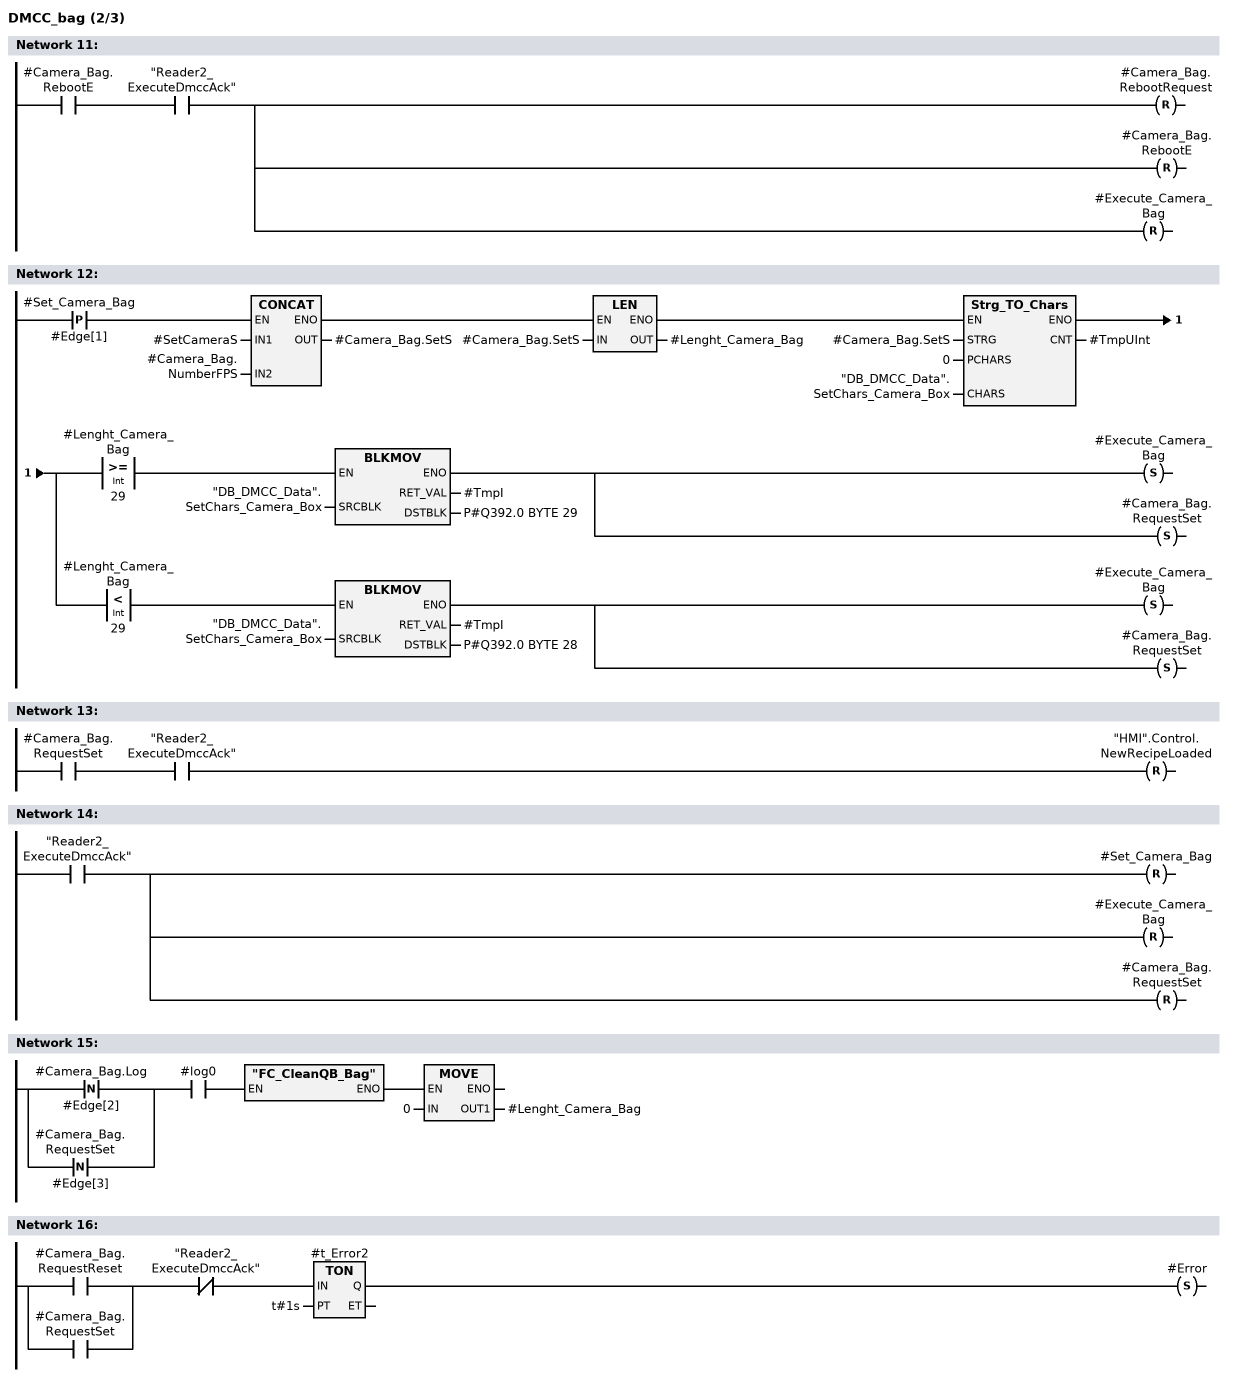
   RUNG wire#powerrail
      Contact( #Camera_Bag.RebootE )
      Contact( "Reader2_ExecuteDmccAck" )
      wire#w1
      R_Coil( #Camera_Bag.RebootRequest )
   END_RUNG
   RUNG wire#w1
      R_Coil( #Camera_Bag.RebootE )
   END_RUNG
   RUNG wire#w1
      R_Coil( #Execute_Camera_Bag )
   END_RUNG
   // the same network as SCL:
   IF #Camera_Bag.RebootE AND "Reader2_ExecuteDmccAck" THEN #Camera_Bag.RebootRequest := FALSE; END_IF;
   #_w1 := #Camera_Bag.RebootE AND "Reader2_ExecuteDmccAck";
   IF #_w1 THEN
       #Camera_Bag.RebootE := FALSE;
       #Execute_Camera_Bag := FALSE;
   END_IF;
END_REGION

REGION Network 12
   // no SCL statement known for Strg_TO_Chars: written as a call
   // ENO of a box is taken as its EN; it also drops when the box reports an error
   #_w1 := #Set_Camera_Bag AND NOT #Edge[1];   // rising edge of #Set_Camera_Bag
   #Edge[1] := #Set_Camera_Bag;
   IF #_w1 THEN
       #Camera_Bag.SetS := CONCAT(IN1 := #SetCameraS, IN2 := #Camera_Bag.NumberFPS);
       #Lenght_Camera_Bag := LEN(IN := #Camera_Bag.SetS);
       Strg_TO_Chars(Strg := #Camera_Bag.SetS,
                     pChars := 0,
                     Chars := "DB_DMCC_Data".SetChars_Camera_Box,
                     Cnt => #TmpUInt);
   END_IF;
   IF #_w1 AND (#Lenght_Camera_Bag >= 29) THEN
       #TmpI := BLKMOV(SRCBLK := "DB_DMCC_Data".SetChars_Camera_Box, DSTBLK => P#Q392.0 BYTE 29);
       #Execute_Camera_Bag := TRUE;
       #Camera_Bag.RequestSet := TRUE;
   END_IF;
   IF #_w1 AND (#Lenght_Camera_Bag < 29) THEN
       #TmpI := BLKMOV(SRCBLK := "DB_DMCC_Data".SetChars_Camera_Box, DSTBLK => P#Q392.0 BYTE 28);
       #Execute_Camera_Bag := TRUE;
       #Camera_Bag.RequestSet := TRUE;
   END_IF;
END_REGION

REGION Network 13
   RUNG wire#powerrail
      Contact( #Camera_Bag.RequestSet )
      Contact( "Reader2_ExecuteDmccAck" )
      R_Coil( "HMI".Control.NewRecipeLoaded )
   END_RUNG
   // the same network as SCL:
   IF #Camera_Bag.RequestSet AND "Reader2_ExecuteDmccAck" THEN
       "HMI".Control.NewRecipeLoaded := FALSE;
   END_IF;
END_REGION

REGION Network 14
   RUNG wire#powerrail
      Contact( "Reader2_ExecuteDmccAck" )
      wire#w1
      R_Coil( #Set_Camera_Bag )
   END_RUNG
   RUNG wire#w1
      R_Coil( #Execute_Camera_Bag )
   END_RUNG
   RUNG wire#w1
      R_Coil( #Camera_Bag.RequestSet )
   END_RUNG
   // the same network as SCL:
   IF "Reader2_ExecuteDmccAck" THEN
       #Set_Camera_Bag := FALSE;
       #Execute_Camera_Bag := FALSE;
       #Camera_Bag.RequestSet := FALSE;
   END_IF;
END_REGION

REGION Network 15
   RUNG wire#powerrail
      N_Contact(operand := #Camera_Bag.Log, bit := #Edge[2])
      wire#w1
      Contact( #log0 )
      "FC_CleanQB_Bag"()
      Move(in := 0, out1 => #Lenght_Camera_Bag)
   END_RUNG
   RUNG wire#powerrail
      N_Contact(operand := #Camera_Bag.RequestSet, bit := #Edge[3])
   END_RUNG wire#w1
   // the same network as SCL:
   #_w1 := NOT #Camera_Bag.Log AND #Edge[2];   // falling edge of #Camera_Bag.Log
   #Edge[2] := #Camera_Bag.Log;
   #_w2 := NOT #Camera_Bag.RequestSet AND #Edge[3];   // falling edge of #Camera_Bag.RequestSet
   #Edge[3] := #Camera_Bag.RequestSet;
   "FC_CleanQB_Bag"(EN := (#_w1 OR #_w2) AND #log0, ENO => #_w3);
   IF #_w3 THEN #Lenght_Camera_Bag := 0; END_IF;
END_REGION

REGION Network 16
   #t_Error2(IN := (#Camera_Bag.RequestReset OR #Camera_Bag.RequestSet) AND NOT "Reader2_ExecuteDmccAck",   // TON
             PT := t#1s);
   IF #t_Error2.Q THEN #Error := TRUE; END_IF;
END_REGION

REGION Network 17
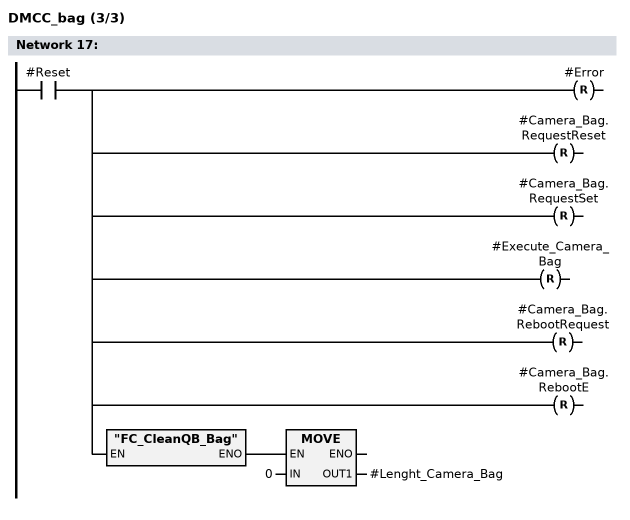
   RUNG wire#powerrail
      Contact( #Reset )
      wire#w1
      R_Coil( #Error )
   END_RUNG
   RUNG wire#w1
      R_Coil( #Camera_Bag.RequestReset )
   END_RUNG
   RUNG wire#w1
      R_Coil( #Camera_Bag.RequestSet )
   END_RUNG
   RUNG wire#w1
      R_Coil( #Execute_Camera_Bag )
   END_RUNG
   RUNG wire#w1
      R_Coil( #Camera_Bag.RebootRequest )
   END_RUNG
   RUNG wire#w1
      R_Coil( #Camera_Bag.RebootE )
   END_RUNG
   RUNG wire#w1
      "FC_CleanQB_Bag"()
      Move(in := 0, out1 => #Lenght_Camera_Bag)
   END_RUNG
   // the same network as SCL:
   IF #Reset THEN
       #Error := FALSE;
       #Camera_Bag.RequestReset := FALSE;
       #Camera_Bag.RequestSet := FALSE;
       #Execute_Camera_Bag := FALSE;
       #Camera_Bag.RebootRequest := FALSE;
       #Camera_Bag.RebootE := FALSE;
   END_IF;
   "FC_CleanQB_Bag"(EN := #Reset, ENO => #_w1);
   IF #_w1 THEN #Lenght_Camera_Bag := 0; END_IF;
END_REGION
END_FUNCTION_BLOCK

FUNCTION_BLOCK "CodeHandle"   // FB105, LAD
{ S7_Optimized_Access := 'TRUE' }
VERSION : 0.1
   VAR_INPUT
      RawCode : Array[0..86] of Char;
      Charakter : String;
      ResultLength : Int;
      Reset_faults : Bool;
      Cam_Box_Read : Bool;
   END_VAR
   VAR_OUTPUT
      LongCode_Out : String[80];
      ShortCode_Out : String[9];
      Read_BOX_EM : Bool;
      Only_ENIGMA : Bool;
      Only_MIRAI : Bool;
   END_VAR
   VAR
      Edge : Array[0..15] of Bool;
      Log1 : Bool;
      Log0 : Bool;
      CharakterPosition : Int;
      RawS : String;
      LongCode : Struct
         Long : String[80];
         Long_Part1 : String[16];
         Long_Part2 : String[12];
         Long_Part3 : String[12];
         Long_Part4 : String[16];
         Long_Part5 : String[8];
         Long_Part6 : String[8];
      END_STRUCT;
      ShortCode : Struct
         ShortCode : String[9];
      END_STRUCT;
      Enigma : TON_TIME;
   END_VAR
   VAR_TEMP
      tmp_w : Word;
      tmp_s : String;
      tmp_small : Bool;
      tmp_big : Bool;
      tmp_read : Bool;
      tmp_read_all : Bool;
   END_VAR
   VAR CONSTANT
      NoCode_ENIGMA : String := 'XXXXXXXXXXXXX';
      NoCode_MIRAI : String := 'XXXXXXXXXXXXXXXXXXXXXXXXXXXXXXXXXXXXXXXXXXXXXXXXXXXXXXXXXXXXXXXXXXXXXX';
   END_VAR
   VAR_TEMP   // added for the SCL form of the ladder/FBD networks
      _w1 : Bool;
      _w2 : Bool;
      _w3 : Bool;
      _w4 : Bool;
      _w5 : Bool;
   END_VAR
BEGIN

REGION Network 1
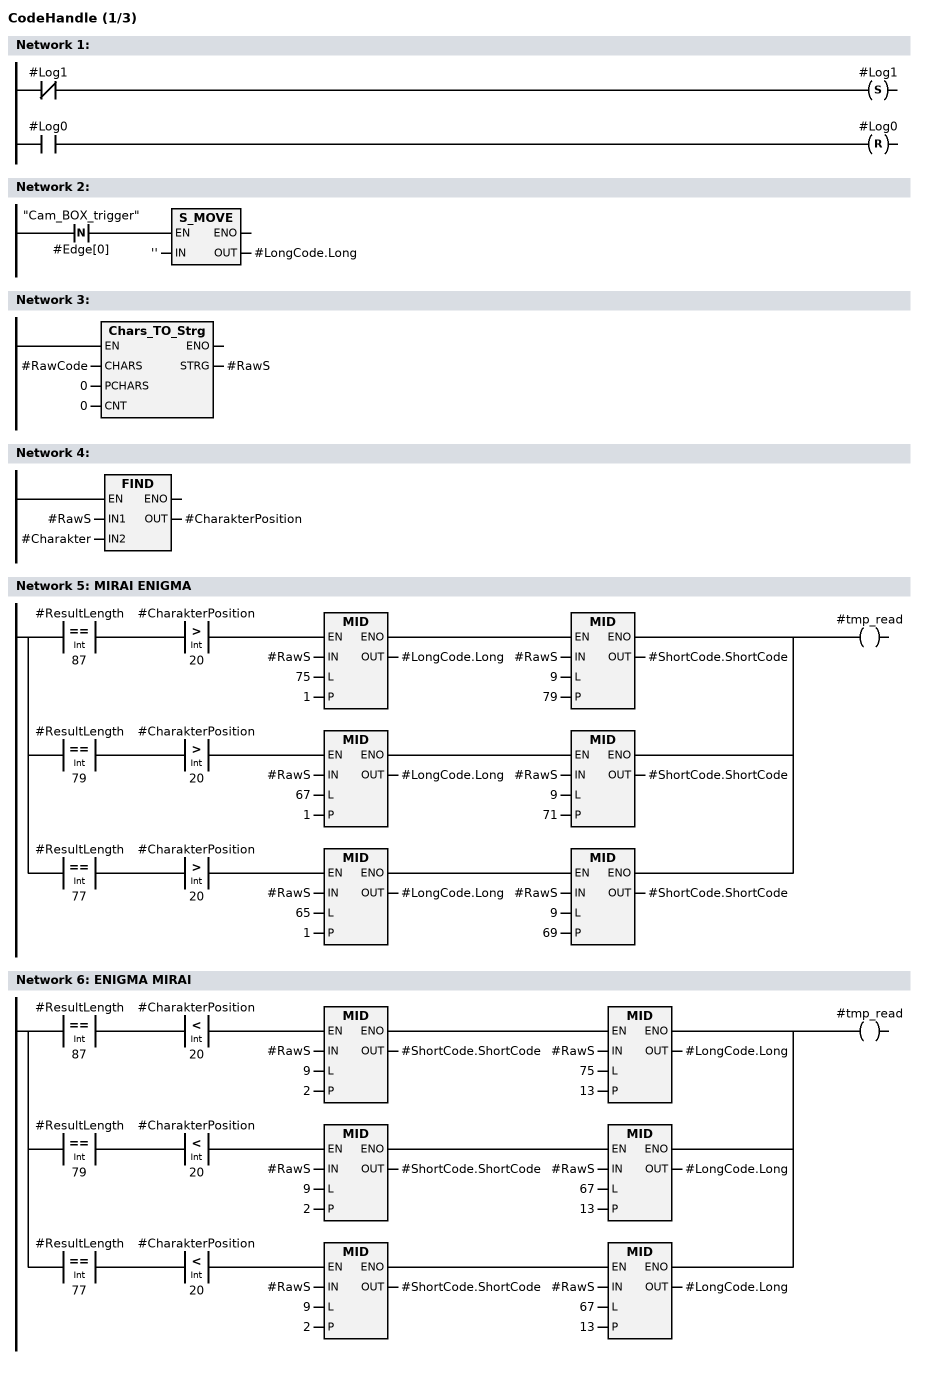
   RUNG wire#powerrail
      I_Contact( #Log1 )
      S_Coil( #Log1 )
   END_RUNG
   RUNG wire#powerrail
      Contact( #Log0 )
      R_Coil( #Log0 )
   END_RUNG
   // the same network as SCL:
   IF NOT #Log1 THEN #Log1 := TRUE; END_IF;
   IF #Log0 THEN #Log0 := FALSE; END_IF;
END_REGION

REGION Network 2
   RUNG wire#powerrail
      N_Contact(operand := "Cam_BOX_trigger", bit := #Edge[0])
      S_Move(in := '', out => #LongCode.Long)
   END_RUNG
   // the same network as SCL:
   #_w1 := NOT "Cam_BOX_trigger" AND #Edge[0];   // falling edge of "Cam_BOX_trigger"
   #Edge[0] := "Cam_BOX_trigger";
   IF #_w1 THEN #LongCode.Long := ''; END_IF;
END_REGION

REGION Network 3
   // no SCL statement known for Chars_TO_Strg: written as a call
   Chars_TO_Strg(Chars := #RawCode, pChars := 0, Cnt := 0, Strg => #RawS);
END_REGION

REGION Network 4
   #CharakterPosition := FIND(IN1 := #RawS, IN2 := #Charakter);
END_REGION

REGION Network 5: MIRAI ENIGMA
   #_w1 := (#ResultLength = 87) AND (#CharakterPosition > 20);
   IF #_w1 THEN
       #LongCode.Long := MID(IN := #RawS, L := 75, P := 1);
       #ShortCode.ShortCode := MID(IN := #RawS, L := 9, P := 79);
   END_IF;
   #_w2 := (#ResultLength = 79) AND (#CharakterPosition > 20);
   IF #_w2 THEN
       #LongCode.Long := MID(IN := #RawS, L := 67, P := 1);
       #ShortCode.ShortCode := MID(IN := #RawS, L := 9, P := 71);
   END_IF;
   #_w3 := (#ResultLength = 77) AND (#CharakterPosition > 20);
   IF #_w3 THEN
       #LongCode.Long := MID(IN := #RawS, L := 65, P := 1);
       #ShortCode.ShortCode := MID(IN := #RawS, L := 9, P := 69);
   END_IF;
   #tmp_read := #_w1 OR #_w2 OR #_w3;
END_REGION

REGION Network 6: ENIGMA MIRAI
   #_w1 := (#ResultLength = 87) AND (#CharakterPosition < 20);
   IF #_w1 THEN
       #ShortCode.ShortCode := MID(IN := #RawS, L := 9, P := 2);
       #LongCode.Long := MID(IN := #RawS, L := 75, P := 13);
   END_IF;
   #_w2 := (#ResultLength = 79) AND (#CharakterPosition < 20);
   IF #_w2 THEN
       #ShortCode.ShortCode := MID(IN := #RawS, L := 9, P := 2);
       #LongCode.Long := MID(IN := #RawS, L := 67, P := 13);
   END_IF;
   #_w3 := (#ResultLength = 77) AND (#CharakterPosition < 20);
   IF #_w3 THEN
       #ShortCode.ShortCode := MID(IN := #RawS, L := 9, P := 2);
       #LongCode.Long := MID(IN := #RawS, L := 67, P := 13);
   END_IF;
   #tmp_read := #_w1 OR #_w2 OR #_w3;
END_REGION

REGION Network 7
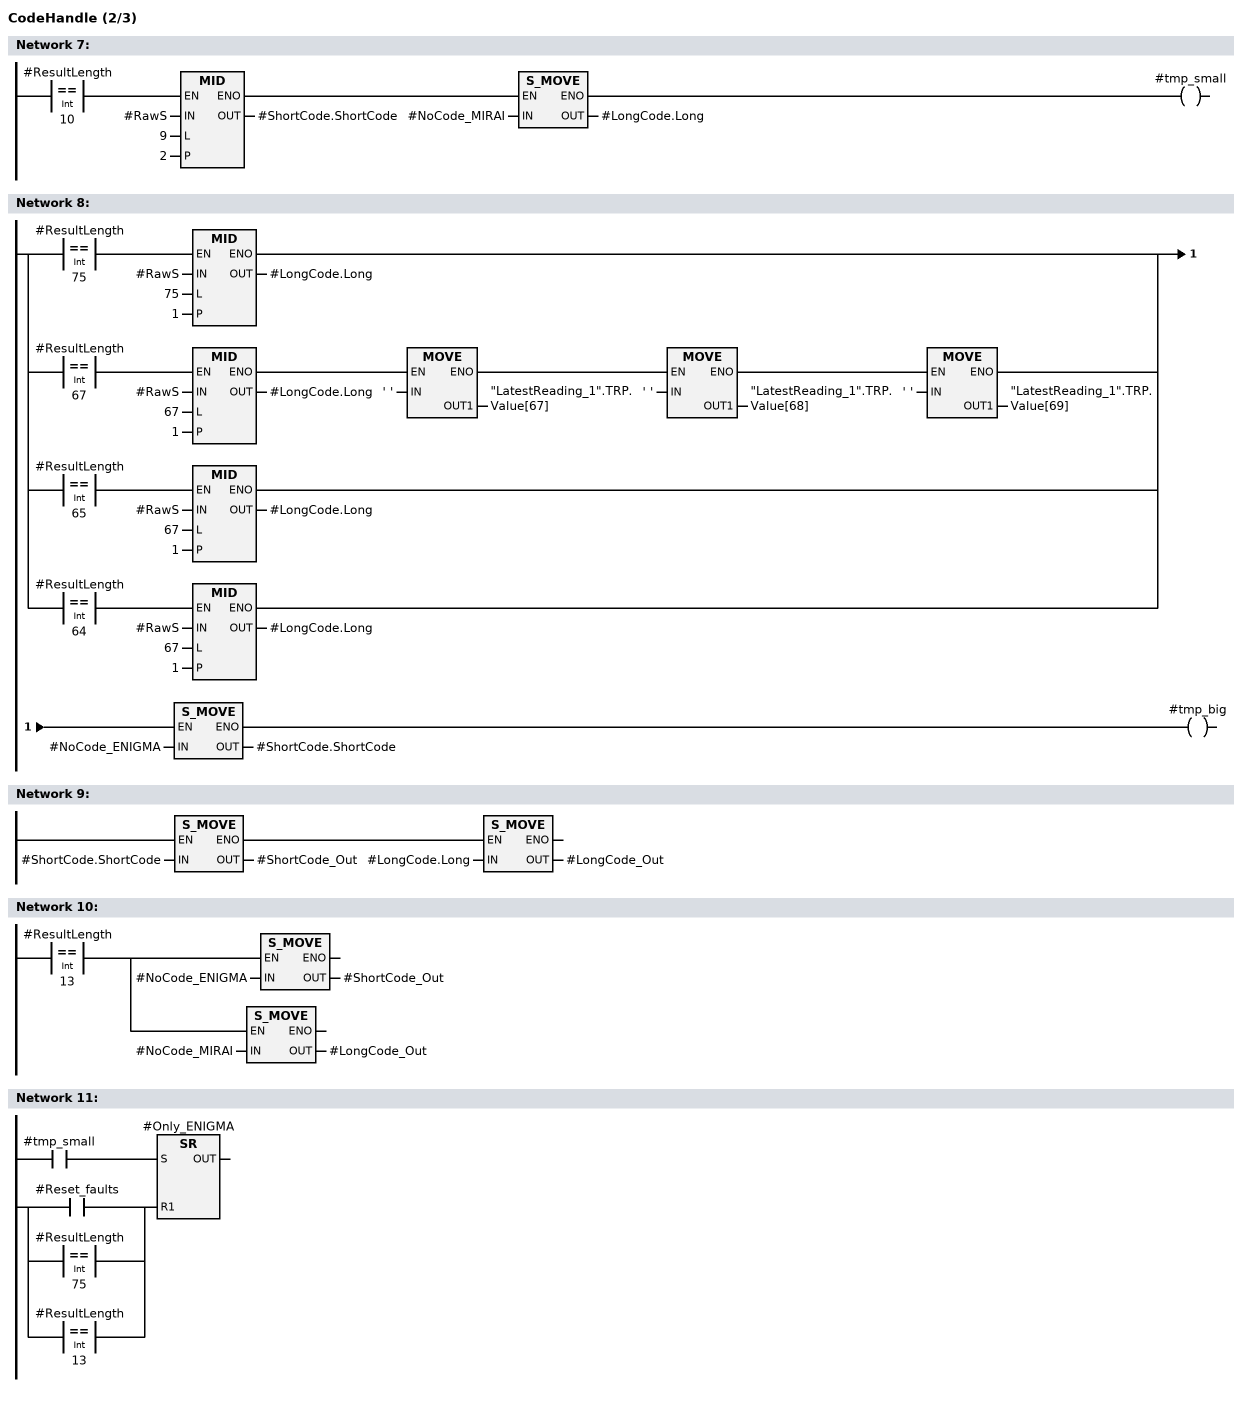
   #_w1 := #ResultLength = 10;
   IF #_w1 THEN
       #ShortCode.ShortCode := MID(IN := #RawS, L := 9, P := 2);
       #LongCode.Long := #NoCode_MIRAI;
   END_IF;
   #tmp_small := #_w1;
END_REGION

REGION Network 8
   #_w1 := #ResultLength = 75;
   IF #_w1 THEN #LongCode.Long := MID(IN := #RawS, L := 75, P := 1); END_IF;
   #_w2 := #ResultLength = 67;
   IF #_w2 THEN
       #LongCode.Long := MID(IN := #RawS, L := 67, P := 1);
       "LatestReading_1".TRP.Value[67] := ' ';
       "LatestReading_1".TRP.Value[68] := ' ';
       "LatestReading_1".TRP.Value[69] := ' ';
   END_IF;
   #_w3 := #ResultLength = 65;
   IF #_w3 THEN #LongCode.Long := MID(IN := #RawS, L := 67, P := 1); END_IF;
   #_w4 := #ResultLength = 64;
   IF #_w4 THEN #LongCode.Long := MID(IN := #RawS, L := 67, P := 1); END_IF;
   #_w5 := #_w1 OR #_w2 OR #_w3 OR #_w4;
   IF #_w5 THEN #ShortCode.ShortCode := #NoCode_ENIGMA; END_IF;
   #tmp_big := #_w5;
END_REGION

REGION Network 9
   RUNG wire#powerrail
      S_Move(in := #ShortCode.ShortCode, out => #ShortCode_Out)
      S_Move(in := #LongCode.Long, out => #LongCode_Out)
   END_RUNG
   // the same network as SCL:
   #ShortCode_Out := #ShortCode.ShortCode;
   #LongCode_Out := #LongCode.Long;
END_REGION

REGION Network 10
   RUNG wire#powerrail
      { S7_Templates := "SrcType := Int" } EQ_Contact(in1 := #ResultLength, in2 := 13)
      wire#w1
      S_Move(in := #NoCode_ENIGMA, out => #ShortCode_Out)
   END_RUNG
   RUNG wire#w1
      S_Move(in := #NoCode_MIRAI, out => #LongCode_Out)
   END_RUNG
   // the same network as SCL:
   IF #ResultLength = 13 THEN
       #ShortCode_Out := #NoCode_ENIGMA;
       #LongCode_Out := #NoCode_MIRAI;
   END_IF;
END_REGION

REGION Network 11
   RUNG wire#powerrail
      Contact( #tmp_small )
      S_SR(operand := #Only_ENIGMA, r1 := wire#w1)
   END_RUNG
   RUNG wire#powerrail
      Contact( #Reset_faults )
   END_RUNG wire#w1
   RUNG wire#powerrail
      { S7_Templates := "SrcType := Int" } EQ_Contact(in1 := #ResultLength, in2 := 75)
   END_RUNG wire#w1
   RUNG wire#powerrail
      { S7_Templates := "SrcType := Int" } EQ_Contact(in1 := #ResultLength, in2 := 13)
   END_RUNG wire#w1
   // the same network as SCL:
   IF #tmp_small THEN
       #Only_ENIGMA := TRUE;   // SR flip-flop
   END_IF;
   IF #Reset_faults OR (#ResultLength = 75) OR (#ResultLength = 13) THEN #Only_ENIGMA := FALSE; END_IF;
END_REGION

REGION Network 12
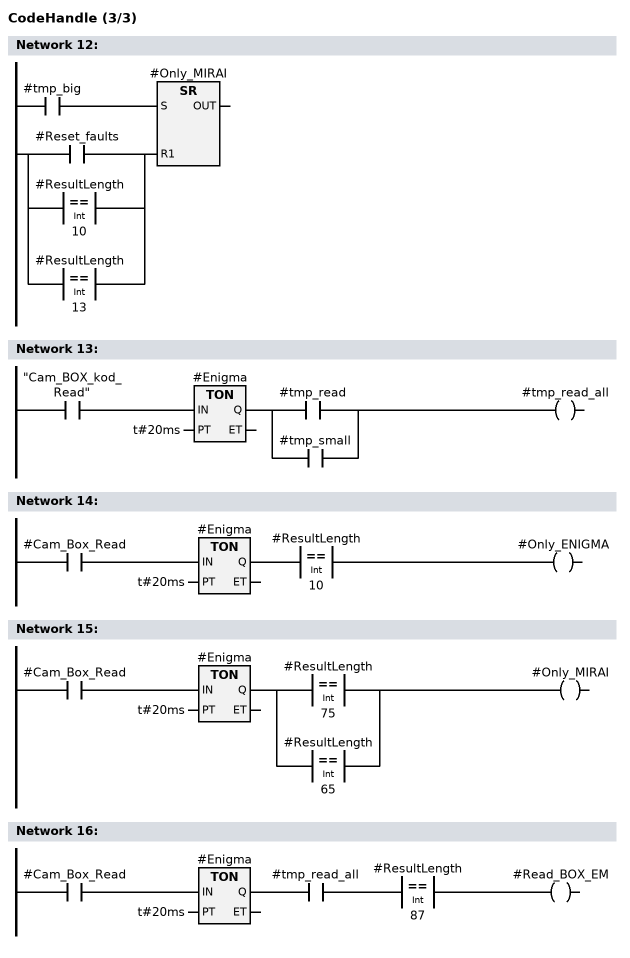
   RUNG wire#powerrail
      Contact( #tmp_big )
      S_SR(operand := #Only_MIRAI, r1 := wire#w1)
   END_RUNG
   RUNG wire#powerrail
      Contact( #Reset_faults )
   END_RUNG wire#w1
   RUNG wire#powerrail
      { S7_Templates := "SrcType := Int" } EQ_Contact(in1 := #ResultLength, in2 := 10)
   END_RUNG wire#w1
   RUNG wire#powerrail
      { S7_Templates := "SrcType := Int" } EQ_Contact(in1 := #ResultLength, in2 := 13)
   END_RUNG wire#w1
   // the same network as SCL:
   IF #tmp_big THEN
       #Only_MIRAI := TRUE;   // SR flip-flop
   END_IF;
   IF #Reset_faults OR (#ResultLength = 10) OR (#ResultLength = 13) THEN #Only_MIRAI := FALSE; END_IF;
END_REGION

REGION Network 13
   #Enigma(IN := "Cam_BOX_kod_Read", PT := t#20ms);   // TON
   #tmp_read_all := #Enigma.Q AND (#tmp_read OR #tmp_small);
END_REGION

REGION Network 14
   #Enigma(IN := #Cam_Box_Read, PT := t#20ms);   // TON
   #Only_ENIGMA := #Enigma.Q AND (#ResultLength = 10);
END_REGION

REGION Network 15
   #Enigma(IN := #Cam_Box_Read, PT := t#20ms);   // TON
   #Only_MIRAI := #Enigma.Q AND ((#ResultLength = 75) OR (#ResultLength = 65));
END_REGION

REGION Network 16
   #Enigma(IN := #Cam_Box_Read, PT := t#20ms);   // TON
   #Read_BOX_EM := #Enigma.Q AND #tmp_read_all AND (#ResultLength = 87);
END_REGION
END_FUNCTION_BLOCK

FUNCTION_BLOCK "LCom_Communication"   // FB30300, SCL
{ S7_Optimized_Access := 'TRUE' }
AUTHOR : APC_ERLF
FAMILY : LCom
VERSION : 2.0
   VAR_INPUT
      enable : Bool := FALSE;
      send : Bool := FALSE;
      sendDataLength : UDInt := 16#FFFFFFFF;
      readDataLength : UDInt := 16#FFFFFFFF;
      configuration : "typeLCom_Config";
   END_VAR
   VAR_OUTPUT
      connected : Bool := FALSE;
      sending : Bool := FALSE;
      dataReceived : Bool := FALSE;
      receivedDataLength : UDInt;
      busy : Bool;
      error : Bool := FALSE;
      status : Word := 16#7000;
   END_VAR
   VAR_IN_OUT
      sendBuffer : Variant;
      receiveBuffer : Variant;
      diagnostics : "typeLCom_Diagnostics";
   END_VAR
   VAR
      statConnectAttempts : SInt;
      statActualLocalLComVersion : USInt;
      statRuntimeTask : LReal;
      statCopyNBytes : UDInt;
      statMaxActPacketLength : UDInt;
      statState : Struct
         connection : USInt := 0;
         cfgSender : USInt;
         comSender : USInt;
         comReceiver : USInt;
         sender : USInt;
         receiver : USInt;
      END_STRUCT;
      statReceive : Struct
         tempTelegram : Struct
            LComVersion : USInt;
            index : USInt;
            telegramType : USInt;
            data : Array[0..23] of Byte;
         END_STRUCT;
         configTelegramV1 : Struct
            LComVersion : USInt;
            telegramType : USInt;
            comMode : USInt;
            slidingWindow : USInt;
            cycleTime : UInt;
            ackTimeOut : UInt;
            lifeSignCycle : UInt;
            status : USInt;
            sendModeSyncTime : USInt;
            maxSendDataLength : UInt;
            maxReceiveDataLength : UInt;
         END_STRUCT;
         configTelegramV2 : Struct
            LComVersion : USInt;
            telegramType : USInt;
            status : USInt;
            sendModeSyncTime : USInt;
            lifeSignCycle : Time;
            cycleTime : Time;
            ackTimeOut : Time;
            maxSendDataLength : UDInt;
            maxReceiveDataLength : UDInt;
         END_STRUCT;
         dataTelegram : Struct
            LComVersion : USInt;
            telegramType : USInt;
            messageCounter : USInt;
            ackMessageCounter : USInt;
            messageOffset : UDInt;
            ackMessageOffset : UDInt;
            actPackageLength : UDInt;
            totalMessageLength : UDInt;
         END_STRUCT;
         userData : Struct
            totalLength : UDInt;
            offset : UDInt;
         END_STRUCT;
         trcvFct : Struct
            data : Array[0..4095] of Byte;
            dataOffset : UDInt;
            dataLength : UDInt;
            dataLengthRest : UDInt;
            dataReceived : Bool := FALSE;
         END_STRUCT;
         numberOfLComHeader : USInt;
      END_STRUCT;
      statSend : Struct
         configTelegramV1 : Struct
            LComVersion : USInt;
            comMode : USInt;
            slidingWindow : USInt;
            cycleTime : UInt;
            ackTimeOut : UInt;
            lifeSignCycle : UInt;
            status : USInt;
            sendModeSyncTime : USInt;
            maxSendDataLength : UInt;
            maxReceiveDataLength : UInt;
         END_STRUCT;
         configTelegramV2 : Struct
            LComVersion : USInt;
            status : USInt;
            sendModeSyncTime : USInt;
            lifeSignCycle : Time;
            cycleTime : Time;
            ackTimeOut : Time;
            maxSendDataLength : UDInt;
            maxReceiveDataLength : UDInt;
         END_STRUCT;
         dataTelegram : Struct
            LComVersion : USInt;
            telegramType : USInt;
            messageCounter : USInt;
            ackMessageCounter : USInt;
            messageOffset : UDInt;
            ackMessageOffset : UDInt;
            actPackageLength : UDInt;
            totalMessageLength : UDInt;
         END_STRUCT;
         userData : Struct
            totalLength : UDInt;
            offset : UDInt;
            sendCycleViolation : Bool;
         END_STRUCT;
         tsendFct : Struct
            dataLengthRest : UInt;
            data : Array[0..4095] of Byte;
            dataOffset : UInt;
            status : Word;
            enable : Bool := FALSE;
         END_STRUCT;
         expectedAck : Struct
            package1 : Struct
               offset : UDInt;
            END_STRUCT;
         END_STRUCT;
         numberOfLComPackage : USInt;
      END_STRUCT;
      statIterator : Int;
      statOldEnable : Bool := FALSE;
      statOldSend : Bool := FALSE;
      statRisingEdgeSend : Bool;
      statFallingEdgeEnable : Bool;
      statRet : Int := -1;
      statCompare : Struct
         sender : Struct
            cycleTime : Time;
            ackTimeOut : Time;
         END_STRUCT;
      END_STRUCT;
      statTconPar : TCON_IP_v4;
      instTCON : TCON;
      instTDISCON : TDISCON;
      instTRCV : TRCV;
      instTSEND : TSEND;
      instLocalLifeSignCycleTimer : TON_TIME;
      instPartnerLifeSignCycleTimer : TON_TIME;
      instLocalCycleTimeTimer : TON_TIME;
      instReceiveMsgCycle : TON_TIME;
      instExpectedAckPackage1 : TON_TIME;
      instMsgSendingTimer : TON_TIME;
      instMsgReceivingTimer : TON_TIME;
      instSyncTimer : TON_TIME;
      instSendErrorTimer : TON_TIME;
      instRcvErrorTimer : TON_TIME;
      instRDREC : RDREC;
      statDiag : Struct
         buffer : Array[0..9] of Struct
            status : Word;
            isActive : Bool;
            subFunctionErrorID : Word;
            additionalValue1 : Real;
            additionalValue2 : Real;
            additionalValue3 : Real;
            additionalValue4 : Time;
         END_STRUCT;
         bufferIndex : USInt := 16#FF;
         actualIndex : USInt;
      END_STRUCT;
   END_VAR
   VAR_TEMP
      tempRuntime : Real;
      tempActTime : DTL;
      tempUDint : UDInt;
      tempDWord : DWord;
   END_VAR
   VAR CONSTANT
      LIFE_SIGN_FACTOR : UInt := 4;
      DIAG_BUFFER_UPPER_LIM : SInt := 63;
      MAX_DATA_BUFFER : Word := 4096;
      LCOM_HEADER_V1 : USInt := 16#10;
      LCOM_HEADER_V2 : USInt := 16#20;
      MAX_TRIAL_TIME : Time := T#200MS;
      STATE_INACTIVE : USInt;
      STATE_INACTIVE_PREPARE : USInt := 1;
      STATE_INIT : USInt := 2;
      OPEN_SERVER : USInt := 3;
      OPEN_CLIENT : USInt := 4;
      OPERATION : USInt := 5;
      FINISH_TSEND : USInt := 6;
      FINISH_TRCV : USInt := 7;
      CALL_TDISCON : USInt := 8;
      CLOSE_CONNECTION : USInt := 9;
      SEND_CONFIG : USInt := 20;
      SEND_DATA : USInt := 30;
      CYCLE : USInt := 31;
      SEND_NO_DATA : USInt := 38;
      NO_CALL_TRCV : USInt := 40;
      READ : USInt := 50;
      NO_DATA_RECEIVED : USInt := 51;
      DATA_RECEIVED : USInt := 52;
      LCOM_EXPECTED : USInt := 53;
      DATA_EXPECTED : USInt := 54;
      WAIT_ACK_TELEGRAM : USInt := 55;
      ACK_TELEGRAM : USInt := 56;
      STATE_WAIT : USInt := 60;
      ERROR_STATE : USInt := 99;
   END_VAR
   // statDiag.buffer[0].isActive := FALSE;
   // statDiag.buffer[1].isActive := FALSE;
   // statDiag.buffer[2].isActive := FALSE;
   // statDiag.buffer[3].isActive := FALSE;
   // statDiag.buffer[4].isActive := FALSE;
   // statDiag.buffer[5].isActive := FALSE;
   // statDiag.buffer[6].isActive := FALSE;
   // statDiag.buffer[7].isActive := FALSE;
   // statDiag.buffer[8].isActive := FALSE;
   // statDiag.buffer[9].isActive := FALSE;
BEGIN
   //=============================================================================
   // SIEMENS AG
   // (c)Copyright 2015 All Rights Reserved
   //-----------------------------------------------------------------------------
   // library: LCom
   // tested with: S7-1215 V4.2, S7-1516 V2.0.1
   // engineering: TIA Portal V14
   // restrictions: none
   // requirements: ---
   // functionality: Function block for TCP communication via Industrial Ethernet.
   // An extended transport protocol, the LCom protocol, has been
   // implemented for extended communication functions.
   // support: profinet.team.motioncontrol.i-dt@siemens.com, Fax: +49(0)9131/98-1297
   // author: APC_ERLF
   //-----------------------------------------------------------------------------
   // change log table:
   // version date        expert in charge changes applied
   // 02.00.03 15.06.2015 APC_ERLF         released version
   // 02.00.04 08.09.2015 APC_ERLF         several bug fixes
   //                                      number of sign-of-life cycles changed from 3 to 4
   // 02.00.05 10.10.2016 APC_ERLF         several bug fixes
   //                                      HW_ANY data type changed (basic data type = UINT)
   //=============================================================================


   //---------------------------------------------------------------------
   //Reset FB outputs, if in the previous cycle are data received
   //---------------------------------------------------------------------
   IF (#dataReceived = TRUE) THEN
     #dataReceived := FALSE;
     #receivedDataLength := 0;

     //Without LCom protocol
     //Leave the FB, if the tcp buffer is not completely analyzed yet
     //Necessary to enforce an L/H edge (FB.dataReceived), if readDataLength is small
     //Example: Rx=100, readDataLength=1
     IF ((NOT #diagnostics.localConfig.connection.useLComProtocol) AND (#statReceive.trcvFct.dataLengthRest > 0)) THEN
       RETURN;
     END_IF;
   END_IF;
   //End:Reset FB outputs, if in the previous cycle data was received


   //---------------------------------------------------------------------
   //Check enable input
   //---------------------------------------------------------------------
   IF ((#enable) AND (NOT #statOldEnable) AND (NOT #statFallingEdgeEnable))//Rising edge
   THEN
     //Start initialize state for the tcp connection
     #statState.connection := #STATE_INIT;
     #status := "LCOM_STATUS_FIRST_CALL";
     #busy := TRUE;
   ELSIF (NOT #enable AND #statState.connection = #STATE_INACTIVE) THEN//Inactive
     RETURN;//Do nothing, wait rising edge on enable
   ELSIF ((NOT #enable) AND (#statOldEnable)) THEN//Falling edge

     #statFallingEdgeEnable := TRUE;
     //LCom Version 1.0 or 2.0 is used OR native tcp
     #statState.connection := #CLOSE_CONNECTION;

     #status := "LCOM_STATUS_DISCONNECTING";
     //Write diagnostics
     #statDiag.bufferIndex := #statDiag.bufferIndex + 1;
     #statDiag.buffer[#statDiag.bufferIndex].#status := "LCOM_STATUS_DISCONNECTING";
     #statDiag.buffer[#statDiag.bufferIndex].subFunctionErrorID := 16#0000;
     #statDiag.buffer[#statDiag.bufferIndex].additionalValue1 := 0.0;
     #statDiag.buffer[#statDiag.bufferIndex].additionalValue2 := 0.0;
     #statDiag.buffer[#statDiag.bufferIndex].additionalValue3 := 0.0;
     #statDiag.buffer[#statDiag.bufferIndex].additionalValue4 := T#0ms;
   ELSE
     ;//No change on enable input
   END_IF;
   #statOldEnable := #enable;
   //End:Check enable input


   // -----------------------------------------------------------------------------------------------------------
   //Statistic --> Calculate average of cycle time [ms]
   // -----------------------------------------------------------------------------------------------------------
   #tempRuntime := (LREAL_TO_REAL(RUNTIME(#statRuntimeTask)) * 1000);

   //Check the measured runtime value and calculate average of cycle time
   IF ((#tempRuntime > 0) AND #enable)
   THEN
     #diagnostics.statistics.avgCallCycle := (((#diagnostics.statistics.avgCallCycle * 49.0) + #tempRuntime) / 50.0);
   ELSE
     ;//Ignore this runtime value 
   END_IF;

   //Initialize values
   #statState.sender := #STATE_INACTIVE;
   #statSend.tsendFct.enable := FALSE;
   #statSend.tsendFct.dataOffset := 0;
   //Set index of temp diagnostics entry
   #statDiag.bufferIndex := 255;
   //End: Calculate average of cycle time and initialize values


   //---------------------------------------------------------------------
   //Check send input
   //---------------------------------------------------------------------
   IF #connected THEN
     //Check rising edge
     IF (#send AND (NOT #statOldSend)) THEN
       //Rising edge detected
       #statRisingEdgeSend := TRUE;
     ELSE
       ;
     END_IF;
     #statOldSend := #send;
   ELSE
     ;//Change at send input is not relevant, because FB is not connected
   END_IF;
   //End:Check send input

   //---------------------------------------------------------------------
   //Acknowledge automatically the followings warnings
   //---------------------------------------------------------------------
   IF (#status = "LCOM_WARN_SEND_DATA_LENGTH")
     OR (#status = "LCOM_WARN_SEND_CYCLE_EXPIRED")
     OR (#status = "LCOM_WARN_RECEIVE_BUFFER_LEN"
     OR (#status = "LCOM_WARN_NO_TIME_SYNC"))
   THEN
     //With LCom protocol
     IF #diagnostics.localConfig.connection.useLComProtocol THEN

       IF (#diagnostics.statistics.activeLComVersion = #LCOM_HEADER_V1) THEN
         #status := "LCOM_STATUS_LCOM_CONNECTED_V1";
       ELSE
         #status := "LCOM_STATUS_LCOM_CONNECTED_V2";
       END_IF;
     ELSE//Without LCom protocol
       #status := "LCOM_STATUS_TCP_CONNECTED";
     END_IF;
   END_IF;
   //End:Acknowledge automatically the followings warnings


   //---------------------------------------------------------------------
   // State machine for IP connection
   //---------------------------------------------------------------------
   CASE #statState.connection OF

     #OPERATION:
       //IP connection is established

       //Get time difference between the last received telegram
       #instPartnerLifeSignCycleTimer(IN := TRUE,
                                      PT := (#diagnostics.partnerConfig.connnection.lifeSignCycleTime * #LIFE_SIGN_FACTOR));

       //Only with LCom protocol, check life sign monitoring
       IF ((#diagnostics.localConfig.connection.useLComProtocol)
         AND
         (#diagnostics.partnerConfig.connnection.lifeSignCycleTime > T#0ms)
         AND
         (#instPartnerLifeSignCycleTimer.Q))
       THEN
         //Write diagnostics
         #statDiag.bufferIndex := #statDiag.bufferIndex + 1;
         #statDiag.buffer[#statDiag.bufferIndex].status := "LCOM_ERR_LIFE_SIGN_EXPIRED";
         #statDiag.buffer[#statDiag.bufferIndex].subFunctionErrorID := 16#0000;
         #statDiag.buffer[#statDiag.bufferIndex].additionalValue1 := UDINT_TO_REAL(TIME_TO_UDINT(#diagnostics.partnerConfig.connnection.lifeSignCycleTime));
         #statDiag.buffer[#statDiag.bufferIndex].additionalValue2 := 0.0;
         #statDiag.buffer[#statDiag.bufferIndex].additionalValue3 := 0.0;
         #statDiag.buffer[#statDiag.bufferIndex].additionalValue4 := #instPartnerLifeSignCycleTimer.ET;

         #statState.connection := #CLOSE_CONNECTION;
         GOTO diag;
       END_IF;

       //---------------------------------------------------------------------
       //Check the status of the "TSEND" instruction of the previous request
       //---------------------------------------------------------------------
       IF ((#statSend.tsendFct.status = 16#7001)
         OR
         (#statSend.tsendFct.status = 16#7002)
         OR
         (#statSend.tsendFct.status = 16#80C4))
       THEN
         //When "TSEND" instruction started or is in sending process
         #instTSEND(REQ := TRUE,
                    LEN := #statSend.tsendFct.dataOffset,
                    ID := #statTconPar.ID,
                    DATA := #statSend.tsendFct.data,
                    STATUS => #statSend.tsendFct.status);

         //When "TSEND" instruction of the previous request is not yet completed
         IF ((#statSend.tsendFct.status = 16#7001)
           OR
           (#statSend.tsendFct.status = 16#7002))
         THEN
           //Stop SendError timer
           #instSendErrorTimer(IN := FALSE,
                               PT := #MAX_TRIAL_TIME);
           RETURN;//"TSEND" instruction still in process, leave FB
         ELSIF (#statSend.tsendFct.status = 16#80C4) THEN
           //Temporary communication error-->Start/Get SendError timer
           #instSendErrorTimer(IN := TRUE,
                               PT := #MAX_TRIAL_TIME);

           //#MAX_TRIAL_TIME is expired
           IF #instSendErrorTimer.Q THEN
             //Write diagnostics
             #statDiag.bufferIndex := #statDiag.bufferIndex + 1;
             #statDiag.buffer[#statDiag.bufferIndex].status := "LCOM_ERR_SEND";
             #statDiag.buffer[#statDiag.bufferIndex].subFunctionErrorID := #statSend.tsendFct.status;
             #statDiag.buffer[#statDiag.bufferIndex].additionalValue1 := 0.0;
             #statDiag.buffer[#statDiag.bufferIndex].additionalValue2 := #statSend.tsendFct.dataOffset;
             #statDiag.buffer[#statDiag.bufferIndex].additionalValue3 := 0.0;
             #statDiag.buffer[#statDiag.bufferIndex].additionalValue4 := T#0ms;
             #statState.connection := #CLOSE_CONNECTION;
             GOTO diag;
           ELSE
             RETURN;//Temporary communication error still valid ant timer is not expired leave FB
           END_IF;
         ELSIF ((#statSend.tsendFct.status = 16#7000) OR (#statSend.tsendFct.status = 16#0000)) THEN
           //---------------------------------------------------------------------
           //Send job completed without error
           //---------------------------------------------------------------------
           IF ((NOT #diagnostics.localConfig.connection.useLComProtocol)
             AND
             (#statSend.userData.offset = #statSend.dataTelegram.totalMessageLength))
           THEN
             //Without LCom protocol
             #statSend.dataTelegram.totalMessageLength := 0;
             #sending := FALSE;

             //Statistic, increase number of sent messages
             #diagnostics.statistics.numberOfSentMessages := #diagnostics.statistics.numberOfSentMessages + 1;

             //Get the message sending time (ms)
             #instMsgSendingTimer(IN := TRUE,
                                  PT := T#+24d20h31m23s647ms);

             //Check maximum message sending time (ms)
             IF (#instMsgSendingTimer.ET > #diagnostics.statistics.maxMsgSendingTime) THEN
               #diagnostics.statistics.maxMsgSendingTime := #instMsgSendingTimer.ET;
             ELSE
               ;//Actual sending time is smaller
             END_IF;

             //Calculate average of message sending time (ms)
             #diagnostics.statistics.avgMsgSendingTime := (((#diagnostics.statistics.avgMsgSendingTime * 19) + UDINT_TO_REAL((TIME_TO_UDINT(#instMsgSendingTimer.ET)))) / 20);